HMI tags "DB_SDC_ERROR_STAT_EMS031"
   "DB_SDC_ERRORS_STAT_ER_AKT[31].ER_TRIGER" : Word = PLC DB_SDC_ERRORS_STAT.ER_AKT[31].ER_TRIGER AT %DB3724.DBW30000, 1 s
   "DB_SDC_ERRORS_STAT_ER_AKT[31].ER_STAT[1].DRIVE_POS" : DInt = PLC DB_SDC_ERRORS_STAT.ER_AKT[31].ER_STAT[1].DRIVE_POS AT %DB3724.DBD30006, 1 s
   "DB_SDC_ERRORS_STAT_ER_AKT[31].ER_STAT[1].ERROR" : Int = PLC DB_SDC_ERRORS_STAT.ER_AKT[31].ER_STAT[1].ERROR AT %DB3724.DBW30012, 1 s
   "DB_SDC_ERRORS_STAT_ER_AKT[31].ER_STAT[2].DRIVE_POS" : DInt = PLC DB_SDC_ERRORS_STAT.ER_AKT[31].ER_STAT[2].DRIVE_POS AT %DB3724.DBD30022, 1 s
   "DB_SDC_ERRORS_STAT_ER_AKT[31].ER_STAT[2].ERROR" : Int = PLC DB_SDC_ERRORS_STAT.ER_AKT[31].ER_STAT[2].ERROR AT %DB3724.DBW30028, 1 s
   "DB_SDC_ERRORS_STAT_ER_AKT[31].ER_STAT[3].DRIVE_POS" : DInt = PLC DB_SDC_ERRORS_STAT.ER_AKT[31].ER_STAT[3].DRIVE_POS AT %DB3724.DBD30038, 1 s
   "DB_SDC_ERRORS_STAT_ER_AKT[31].ER_STAT[3].ERROR" : Int = PLC DB_SDC_ERRORS_STAT.ER_AKT[31].ER_STAT[3].ERROR AT %DB3724.DBW30044, 1 s
   "DB_SDC_ERRORS_STAT_ER_AKT[31].ER_STAT[4].DRIVE_POS" : DInt = PLC DB_SDC_ERRORS_STAT.ER_AKT[31].ER_STAT[4].DRIVE_POS AT %DB3724.DBD30054, 1 s
   "DB_SDC_ERRORS_STAT_ER_AKT[31].ER_STAT[4].ERROR" : Int = PLC DB_SDC_ERRORS_STAT.ER_AKT[31].ER_STAT[4].ERROR AT %DB3724.DBW30060, 1 s

HMI tags "DB_SDC_ERROR_STAT_EMS032"
   "DB_SDC_ERRORS_STAT_ER_AKT[32].ER_TRIGER" : Word = PLC DB_SDC_ERRORS_STAT.ER_AKT[32].ER_TRIGER AT %DB3724.DBW30066, 1 s
   "DB_SDC_ERRORS_STAT_ER_AKT[32].ER_STAT[1].DRIVE_POS" : DInt = PLC DB_SDC_ERRORS_STAT.ER_AKT[32].ER_STAT[1].DRIVE_POS AT %DB3724.DBD30072, 1 s
   "DB_SDC_ERRORS_STAT_ER_AKT[32].ER_STAT[1].ERROR" : Int = PLC DB_SDC_ERRORS_STAT.ER_AKT[32].ER_STAT[1].ERROR AT %DB3724.DBW30078, 1 s
   "DB_SDC_ERRORS_STAT_ER_AKT[32].ER_STAT[2].DRIVE_POS" : DInt = PLC DB_SDC_ERRORS_STAT.ER_AKT[32].ER_STAT[2].DRIVE_POS AT %DB3724.DBD30088, 1 s
   "DB_SDC_ERRORS_STAT_ER_AKT[32].ER_STAT[2].ERROR" : Int = PLC DB_SDC_ERRORS_STAT.ER_AKT[32].ER_STAT[2].ERROR AT %DB3724.DBW30094, 1 s
   "DB_SDC_ERRORS_STAT_ER_AKT[32].ER_STAT[3].DRIVE_POS" : DInt = PLC DB_SDC_ERRORS_STAT.ER_AKT[32].ER_STAT[3].DRIVE_POS AT %DB3724.DBD30104, 1 s
   "DB_SDC_ERRORS_STAT_ER_AKT[32].ER_STAT[3].ERROR" : Int = PLC DB_SDC_ERRORS_STAT.ER_AKT[32].ER_STAT[3].ERROR AT %DB3724.DBW30110, 1 s
   "DB_SDC_ERRORS_STAT_ER_AKT[32].ER_STAT[4].DRIVE_POS" : DInt = PLC DB_SDC_ERRORS_STAT.ER_AKT[32].ER_STAT[4].DRIVE_POS AT %DB3724.DBD30120, 1 s
   "DB_SDC_ERRORS_STAT_ER_AKT[32].ER_STAT[4].ERROR" : Int = PLC DB_SDC_ERRORS_STAT.ER_AKT[32].ER_STAT[4].ERROR AT %DB3724.DBW30126, 1 s

HMI tags "DB_SDC_ERROR_STAT_EMS033"
   "DB_SDC_ERRORS_STAT_ER_AKT[33].ER_TRIGER" : Word = PLC DB_SDC_ERRORS_STAT.ER_AKT[33].ER_TRIGER AT %DB3724.DBW30132, 1 s
   "DB_SDC_ERRORS_STAT_ER_AKT[33].ER_STAT[1].DRIVE_POS" : DInt = PLC DB_SDC_ERRORS_STAT.ER_AKT[33].ER_STAT[1].DRIVE_POS AT %DB3724.DBD30138, 1 s
   "DB_SDC_ERRORS_STAT_ER_AKT[33].ER_STAT[1].ERROR" : Int = PLC DB_SDC_ERRORS_STAT.ER_AKT[33].ER_STAT[1].ERROR AT %DB3724.DBW30144, 1 s
   "DB_SDC_ERRORS_STAT_ER_AKT[33].ER_STAT[2].DRIVE_POS" : DInt = PLC DB_SDC_ERRORS_STAT.ER_AKT[63].ER_STAT[4].DRIVE_POS AT %DB3724.DBD30154, 1 s
   "DB_SDC_ERRORS_STAT_ER_AKT[33].ER_STAT[2].ERROR" : Int = PLC DB_SDC_ERRORS_STAT.ER_AKT[33].ER_STAT[2].ERROR AT %DB3724.DBW30160, 1 s
   "DB_SDC_ERRORS_STAT_ER_AKT[33].ER_STAT[3].DRIVE_POS" : DInt = PLC DB_SDC_ERRORS_STAT.ER_AKT[33].ER_STAT[3].DRIVE_POS AT %DB3724.DBD30170, 1 s
   "DB_SDC_ERRORS_STAT_ER_AKT[33].ER_STAT[3].ERROR" : Int = PLC DB_SDC_ERRORS_STAT.ER_AKT[33].ER_STAT[3].ERROR AT %DB3724.DBW30176, 1 s
   "DB_SDC_ERRORS_STAT_ER_AKT[33].ER_STAT[4].DRIVE_POS" : DInt = PLC DB_SDC_ERRORS_STAT.ER_AKT[33].ER_STAT[4].DRIVE_POS AT %DB3724.DBD30186, 1 s
   "DB_SDC_ERRORS_STAT_ER_AKT[33].ER_STAT[4].ERROR" : Int = PLC DB_SDC_ERRORS_STAT.ER_AKT[33].ER_STAT[4].ERROR AT %DB3724.DBW30192, 1 s

HMI tags "DB_SDC_ERROR_STAT_EMS034"
   "DB_SDC_ERRORS_STAT_ER_AKT[34].ER_TRIGER" : Word = PLC DB_SDC_ERRORS_STAT.ER_AKT[34].ER_TRIGER AT %DB3724.DBW30198, 1 s
   "DB_SDC_ERRORS_STAT_ER_AKT[34].ER_STAT[1].DRIVE_POS" : DInt = PLC DB_SDC_ERRORS_STAT.ER_AKT[34].ER_STAT[1].DRIVE_POS AT %DB3724.DBD30204, 1 s
   "DB_SDC_ERRORS_STAT_ER_AKT[34].ER_STAT[1].ERROR" : Int = PLC DB_SDC_ERRORS_STAT.ER_AKT[34].ER_STAT[1].ERROR AT %DB3724.DBW30210, 1 s
   "DB_SDC_ERRORS_STAT_ER_AKT[34].ER_STAT[2].DRIVE_POS" : DInt = PLC DB_SDC_ERRORS_STAT.ER_AKT[34].ER_STAT[2].DRIVE_POS AT %DB3724.DBD30220, 1 s
   "DB_SDC_ERRORS_STAT_ER_AKT[34].ER_STAT[2].ERROR" : Int = PLC DB_SDC_ERRORS_STAT.ER_AKT[34].ER_STAT[2].ERROR AT %DB3724.DBW30226, 1 s
   "DB_SDC_ERRORS_STAT_ER_AKT[34].ER_STAT[3].DRIVE_POS" : DInt = PLC DB_SDC_ERRORS_STAT.ER_AKT[34].ER_STAT[3].DRIVE_POS AT %DB3724.DBD30236, 1 s
   "DB_SDC_ERRORS_STAT_ER_AKT[34].ER_STAT[3].ERROR" : Int = PLC DB_SDC_ERRORS_STAT.ER_AKT[34].ER_STAT[3].ERROR AT %DB3724.DBW30242, 1 s
   "DB_SDC_ERRORS_STAT_ER_AKT[34].ER_STAT[4].DRIVE_POS" : DInt = PLC DB_SDC_ERRORS_STAT.ER_AKT[34].ER_STAT[4].DRIVE_POS AT %DB3724.DBD30252, 1 s
   "DB_SDC_ERRORS_STAT_ER_AKT[34].ER_STAT[4].ERROR" : Int = PLC DB_SDC_ERRORS_STAT.ER_AKT[34].ER_STAT[4].ERROR AT %DB3724.DBW30258, 1 s

HMI tags "DB_SDC_ERROR_STAT_EMS035"
   "DB_SDC_ERRORS_STAT_ER_AKT[35].ER_TRIGER" : Word = PLC DB_SDC_ERRORS_STAT.ER_AKT[35].ER_TRIGER AT %DB3724.DBW30264, 1 s
   "DB_SDC_ERRORS_STAT_ER_AKT[35].ER_STAT[1].DRIVE_POS" : DInt = PLC DB_SDC_ERRORS_STAT.ER_AKT[35].ER_STAT[1].DRIVE_POS AT %DB3724.DBD30270, 1 s
   "DB_SDC_ERRORS_STAT_ER_AKT[35].ER_STAT[1].ERROR" : Int = PLC DB_SDC_ERRORS_STAT.ER_AKT[35].ER_STAT[1].ERROR AT %DB3724.DBW30276, 1 s
   "DB_SDC_ERRORS_STAT_ER_AKT[35].ER_STAT[2].DRIVE_POS" : DInt = PLC DB_SDC_ERRORS_STAT.ER_AKT[35].ER_STAT[2].DRIVE_POS AT %DB3724.DBD30286, 1 s
   "DB_SDC_ERRORS_STAT_ER_AKT[35].ER_STAT[2].ERROR" : Int = PLC DB_SDC_ERRORS_STAT.ER_AKT[35].ER_STAT[2].ERROR AT %DB3724.DBW30292, 1 s
   "DB_SDC_ERRORS_STAT_ER_AKT[35].ER_STAT[3].DRIVE_POS" : DInt = PLC DB_SDC_ERRORS_STAT.ER_AKT[35].ER_STAT[3].DRIVE_POS AT %DB3724.DBD30302, 1 s
   "DB_SDC_ERRORS_STAT_ER_AKT[35].ER_STAT[3].ERROR" : Int = PLC DB_SDC_ERRORS_STAT.ER_AKT[35].ER_STAT[3].ERROR AT %DB3724.DBW30308, 1 s
   "DB_SDC_ERRORS_STAT_ER_AKT[35].ER_STAT[4].DRIVE_POS" : DInt = PLC DB_SDC_ERRORS_STAT.ER_AKT[35].ER_STAT[4].DRIVE_POS AT %DB3724.DBD30318, 1 s
   "DB_SDC_ERRORS_STAT_ER_AKT[35].ER_STAT[4].ERROR" : Int = PLC DB_SDC_ERRORS_STAT.ER_AKT[35].ER_STAT[4].ERROR AT %DB3724.DBW30324, 1 s

HMI tags "DB_SDC_ERROR_STAT_EMS036"
   "DB_SDC_ERRORS_STAT_ER_AKT[36].ER_TRIGER" : Word = PLC DB_SDC_ERRORS_STAT.ER_AKT[36].ER_TRIGER AT %DB3724.DBW30330, 1 s
   "DB_SDC_ERRORS_STAT_ER_AKT[36].ER_STAT[1].DRIVE_POS" : DInt = PLC DB_SDC_ERRORS_STAT.ER_AKT[36].ER_STAT[1].DRIVE_POS AT %DB3724.DBD30336, 1 s
   "DB_SDC_ERRORS_STAT_ER_AKT[36].ER_STAT[1].ERROR" : Int = PLC DB_SDC_ERRORS_STAT.ER_AKT[36].ER_STAT[1].ERROR AT %DB3724.DBW30342, 1 s
   "DB_SDC_ERRORS_STAT_ER_AKT[36].ER_STAT[2].DRIVE_POS" : DInt = PLC DB_SDC_ERRORS_STAT.ER_AKT[36].ER_STAT[2].DRIVE_POS AT %DB3724.DBD30352, 1 s
   "DB_SDC_ERRORS_STAT_ER_AKT[36].ER_STAT[2].ERROR" : Int = PLC DB_SDC_ERRORS_STAT.ER_AKT[36].ER_STAT[2].ERROR AT %DB3724.DBW30358, 1 s
   "DB_SDC_ERRORS_STAT_ER_AKT[36].ER_STAT[3].DRIVE_POS" : DInt = PLC DB_SDC_ERRORS_STAT.ER_AKT[36].ER_STAT[3].DRIVE_POS AT %DB3724.DBD30368, 1 s
   "DB_SDC_ERRORS_STAT_ER_AKT[36].ER_STAT[3].ERROR" : Int = PLC DB_SDC_ERRORS_STAT.ER_AKT[36].ER_STAT[3].ERROR AT %DB3724.DBW30374, 1 s
   "DB_SDC_ERRORS_STAT_ER_AKT[36].ER_STAT[4].DRIVE_POS" : DInt = PLC DB_SDC_ERRORS_STAT.ER_AKT[36].ER_STAT[4].DRIVE_POS AT %DB3724.DBD30384, 1 s
   "DB_SDC_ERRORS_STAT_ER_AKT[36].ER_STAT[4].ERROR" : Int = PLC DB_SDC_ERRORS_STAT.ER_AKT[36].ER_STAT[4].ERROR AT %DB3724.DBW30390, 1 s

HMI tags "DB_SDC_ERROR_STAT_EMS037"
   "DB_SDC_ERRORS_STAT_ER_AKT[37].ER_TRIGER" : Word = PLC DB_SDC_ERRORS_STAT.ER_AKT[37].ER_TRIGER AT %DB3724.DBW30396, 1 s
   "DB_SDC_ERRORS_STAT_ER_AKT[37].ER_STAT[1].DRIVE_POS" : DInt = PLC DB_SDC_ERRORS_STAT.ER_AKT[37].ER_STAT[1].DRIVE_POS AT %DB3724.DBD30402, 1 s
   "DB_SDC_ERRORS_STAT_ER_AKT[37].ER_STAT[1].ERROR" : Int = PLC DB_SDC_ERRORS_STAT.ER_AKT[37].ER_STAT[1].ERROR AT %DB3724.DBW30408, 1 s
   "DB_SDC_ERRORS_STAT_ER_AKT[37].ER_STAT[2].DRIVE_POS" : DInt = PLC DB_SDC_ERRORS_STAT.ER_AKT[37].ER_STAT[2].DRIVE_POS AT %DB3724.DBD30418, 1 s
   "DB_SDC_ERRORS_STAT_ER_AKT[37].ER_STAT[2].ERROR" : Int = PLC DB_SDC_ERRORS_STAT.ER_AKT[37].ER_STAT[2].ERROR AT %DB3724.DBW30424, 1 s
   "DB_SDC_ERRORS_STAT_ER_AKT[37].ER_STAT[3].DRIVE_POS" : DInt = PLC DB_SDC_ERRORS_STAT.ER_AKT[37].ER_STAT[3].DRIVE_POS AT %DB3724.DBD30434, 1 s
   "DB_SDC_ERRORS_STAT_ER_AKT[37].ER_STAT[3].ERROR" : Int = PLC DB_SDC_ERRORS_STAT.ER_AKT[37].ER_STAT[3].ERROR AT %DB3724.DBW30440, 1 s
   "DB_SDC_ERRORS_STAT_ER_AKT[37].ER_STAT[4].DRIVE_POS" : DInt = PLC DB_SDC_ERRORS_STAT.ER_AKT[37].ER_STAT[4].DRIVE_POS AT %DB3724.DBD30450, 1 s
   "DB_SDC_ERRORS_STAT_ER_AKT[37].ER_STAT[4].ERROR" : Int = PLC DB_SDC_ERRORS_STAT.ER_AKT[37].ER_STAT[4].ERROR AT %DB3724.DBW30456, 1 s

HMI tags "DB_SDC_ERROR_STAT_EMS038"
   "DB_SDC_ERRORS_STAT_ER_AKT[38].ER_TRIGER" : Word = PLC DB_SDC_ERRORS_STAT.ER_AKT[38].ER_TRIGER AT %DB3724.DBW30462, 1 s
   "DB_SDC_ERRORS_STAT_ER_AKT[38].ER_STAT[1].DRIVE_POS" : DInt = PLC DB_SDC_ERRORS_STAT.ER_AKT[38].ER_STAT[1].DRIVE_POS AT %DB3724.DBD30468, 1 s
   "DB_SDC_ERRORS_STAT_ER_AKT[38].ER_STAT[1].ERROR" : Int = PLC DB_SDC_ERRORS_STAT.ER_AKT[38].ER_STAT[1].ERROR AT %DB3724.DBW30474, 1 s
   "DB_SDC_ERRORS_STAT_ER_AKT[38].ER_STAT[2].DRIVE_POS" : DInt = PLC DB_SDC_ERRORS_STAT.ER_AKT[38].ER_STAT[2].DRIVE_POS AT %DB3724.DBD30484, 1 s
   "DB_SDC_ERRORS_STAT_ER_AKT[38].ER_STAT[2].ERROR" : Int = PLC DB_SDC_ERRORS_STAT.ER_AKT[38].ER_STAT[2].ERROR AT %DB3724.DBW30490, 1 s
   "DB_SDC_ERRORS_STAT_ER_AKT[38].ER_STAT[3].DRIVE_POS" : DInt = PLC DB_SDC_ERRORS_STAT.ER_AKT[38].ER_STAT[3].DRIVE_POS AT %DB3724.DBD30500, 1 s
   "DB_SDC_ERRORS_STAT_ER_AKT[38].ER_STAT[3].ERROR" : Int = PLC DB_SDC_ERRORS_STAT.ER_AKT[38].ER_STAT[3].ERROR AT %DB3724.DBW30506, 1 s
   "DB_SDC_ERRORS_STAT_ER_AKT[38].ER_STAT[4].DRIVE_POS" : DInt = PLC DB_SDC_ERRORS_STAT.ER_AKT[38].ER_STAT[4].DRIVE_POS AT %DB3724.DBD30516, 1 s
   "DB_SDC_ERRORS_STAT_ER_AKT[38].ER_STAT[4].ERROR" : Int = PLC DB_SDC_ERRORS_STAT.ER_AKT[38].ER_STAT[4].ERROR AT %DB3724.DBW30522, 1 s

HMI tags "DB_SDC_ERROR_STAT_EMS039"
   "DB_SDC_ERRORS_STAT_ER_AKT[39].ER_TRIGER" : Word = PLC DB_SDC_ERRORS_STAT.ER_AKT[39].ER_TRIGER AT %DB3724.DBW30528, 1 s
   "DB_SDC_ERRORS_STAT_ER_AKT[39].ER_STAT[1].DRIVE_POS" : DInt = PLC DB_SDC_ERRORS_STAT.ER_AKT[39].ER_STAT[1].DRIVE_POS AT %DB3724.DBD30534, 1 s
   "DB_SDC_ERRORS_STAT_ER_AKT[39].ER_STAT[1].ERROR" : Int = PLC DB_SDC_ERRORS_STAT.ER_AKT[39].ER_STAT[1].ERROR AT %DB3724.DBW30540, 1 s
   "DB_SDC_ERRORS_STAT_ER_AKT[39].ER_STAT[2].DRIVE_POS" : DInt = PLC DB_SDC_ERRORS_STAT.ER_AKT[39].ER_STAT[2].DRIVE_POS AT %DB3724.DBD30550, 1 s
   "DB_SDC_ERRORS_STAT_ER_AKT[39].ER_STAT[2].ERROR" : Int = PLC DB_SDC_ERRORS_STAT.ER_AKT[39].ER_STAT[2].ERROR AT %DB3724.DBW30556, 1 s
   "DB_SDC_ERRORS_STAT_ER_AKT[39].ER_STAT[3].DRIVE_POS" : DInt = PLC DB_SDC_ERRORS_STAT.ER_AKT[39].ER_STAT[3].DRIVE_POS AT %DB3724.DBD30566, 1 s
   "DB_SDC_ERRORS_STAT_ER_AKT[39].ER_STAT[3].ERROR" : Int = PLC DB_SDC_ERRORS_STAT.ER_AKT[39].ER_STAT[3].ERROR AT %DB3724.DBW30572, 1 s
   "DB_SDC_ERRORS_STAT_ER_AKT[39].ER_STAT[4].DRIVE_POS" : DInt = PLC DB_SDC_ERRORS_STAT.ER_AKT[39].ER_STAT[4].DRIVE_POS AT %DB3724.DBD30582, 1 s
   "DB_SDC_ERRORS_STAT_ER_AKT[39].ER_STAT[4].ERROR" : Int = PLC DB_SDC_ERRORS_STAT.ER_AKT[39].ER_STAT[4].ERROR AT %DB3724.DBW30588, 1 s

HMI tags "DB_SDC_ERROR_STAT_EMS040"
   "DB_SDC_ERRORS_STAT_ER_AKT[40].ER_TRIGER" : Word = PLC DB_SDC_ERRORS_STAT.ER_AKT[40].ER_TRIGER AT %DB3724.DBW30594, 1 s
   "DB_SDC_ERRORS_STAT_ER_AKT[40].ER_STAT[1].DRIVE_POS" : DInt = PLC DB_SDC_ERRORS_STAT.ER_AKT[40].ER_STAT[1].DRIVE_POS AT %DB3724.DBD30600, 1 s
   "DB_SDC_ERRORS_STAT_ER_AKT[40].ER_STAT[1].ERROR" : Int = PLC DB_SDC_ERRORS_STAT.ER_AKT[40].ER_STAT[1].ERROR AT %DB3724.DBW30606, 1 s
   "DB_SDC_ERRORS_STAT_ER_AKT[40].ER_STAT[2].DRIVE_POS" : DInt = PLC DB_SDC_ERRORS_STAT.ER_AKT[40].ER_STAT[2].DRIVE_POS AT %DB3724.DBD30616, 1 s
   "DB_SDC_ERRORS_STAT_ER_AKT[40].ER_STAT[2].ERROR" : Int = PLC DB_SDC_ERRORS_STAT.ER_AKT[40].ER_STAT[2].ERROR AT %DB3724.DBW30622, 1 s
   "DB_SDC_ERRORS_STAT_ER_AKT[40].ER_STAT[3].DRIVE_POS" : DInt = PLC DB_SDC_ERRORS_STAT.ER_AKT[40].ER_STAT[3].DRIVE_POS AT %DB3724.DBD30632, 1 s
   "DB_SDC_ERRORS_STAT_ER_AKT[40].ER_STAT[3].ERROR" : Int = PLC DB_SDC_ERRORS_STAT.ER_AKT[40].ER_STAT[3].ERROR AT %DB3724.DBW30638, 1 s
   "DB_SDC_ERRORS_STAT_ER_AKT[40].ER_STAT[4].DRIVE_POS" : DInt = PLC DB_SDC_ERRORS_STAT.ER_AKT[40].ER_STAT[4].DRIVE_POS AT %DB3724.DBD30648, 1 s
   "DB_SDC_ERRORS_STAT_ER_AKT[40].ER_STAT[4].ERROR" : Int = PLC DB_SDC_ERRORS_STAT.ER_AKT[40].ER_STAT[4].ERROR AT %DB3724.DBW30654, 1 s

HMI tags "DB_SDC_ERROR_STAT_EMS041"
   "DB_SDC_ERRORS_STAT_ER_AKT[41].ER_TRIGER" : Word = PLC DB_SDC_ERRORS_STAT.ER_AKT[41].ER_TRIGER AT %DB3724.DBW30660, 1 s
   "DB_SDC_ERRORS_STAT_ER_AKT[41].ER_STAT[1].DRIVE_POS" : DInt = PLC DB_SDC_ERRORS_STAT.ER_AKT[41].ER_STAT[1].DRIVE_POS AT %DB3724.DBD30666, 1 s
   "DB_SDC_ERRORS_STAT_ER_AKT[41].ER_STAT[1].ERROR" : Int = PLC DB_SDC_ERRORS_STAT.ER_AKT[41].ER_STAT[1].ERROR AT %DB3724.DBW30672, 1 s
   "DB_SDC_ERRORS_STAT_ER_AKT[41].ER_STAT[2].DRIVE_POS" : DInt = PLC DB_SDC_ERRORS_STAT.ER_AKT[41].ER_STAT[2].DRIVE_POS AT %DB3724.DBD30682, 1 s
   "DB_SDC_ERRORS_STAT_ER_AKT[41].ER_STAT[2].ERROR" : Int = PLC DB_SDC_ERRORS_STAT.ER_AKT[41].ER_STAT[2].ERROR AT %DB3724.DBW30688, 1 s
   "DB_SDC_ERRORS_STAT_ER_AKT[41].ER_STAT[3].DRIVE_POS" : DInt = PLC DB_SDC_ERRORS_STAT.ER_AKT[41].ER_STAT[3].DRIVE_POS AT %DB3724.DBD30698, 1 s
   "DB_SDC_ERRORS_STAT_ER_AKT[41].ER_STAT[3].ERROR" : Int = PLC DB_SDC_ERRORS_STAT.ER_AKT[41].ER_STAT[3].ERROR AT %DB3724.DBW30704, 1 s
   "DB_SDC_ERRORS_STAT_ER_AKT[41].ER_STAT[4].DRIVE_POS" : DInt = PLC DB_SDC_ERRORS_STAT.ER_AKT[41].ER_STAT[4].DRIVE_POS AT %DB3724.DBD30714, 1 s
   "DB_SDC_ERRORS_STAT_ER_AKT[41].ER_STAT[4].ERROR" : Int = PLC DB_SDC_ERRORS_STAT.ER_AKT[41].ER_STAT[4].ERROR AT %DB3724.DBW30720, 1 s

HMI tags "DB_SDC_ERROR_STAT_EMS042"
   "DB_SDC_ERRORS_STAT_ER_AKT[42].ER_TRIGER" : Word = PLC DB_SDC_ERRORS_STAT.ER_AKT[42].ER_TRIGER AT %DB3724.DBW30726, 1 s
   "DB_SDC_ERRORS_STAT_ER_AKT[42].ER_STAT[1].DRIVE_POS" : DInt = PLC DB_SDC_ERRORS_STAT.ER_AKT[42].ER_STAT[1].DRIVE_POS AT %DB3724.DBD30732, 1 s
   "DB_SDC_ERRORS_STAT_ER_AKT[42].ER_STAT[1].ERROR" : Int = PLC DB_SDC_ERRORS_STAT.ER_AKT[42].ER_STAT[1].ERROR AT %DB3724.DBW30738, 1 s
   "DB_SDC_ERRORS_STAT_ER_AKT[42].ER_STAT[2].DRIVE_POS" : DInt = PLC DB_SDC_ERRORS_STAT.ER_AKT[42].ER_STAT[2].DRIVE_POS AT %DB3724.DBD30748, 1 s
   "DB_SDC_ERRORS_STAT_ER_AKT[42].ER_STAT[2].ERROR" : Int = PLC DB_SDC_ERRORS_STAT.ER_AKT[42].ER_STAT[2].ERROR AT %DB3724.DBW30754, 1 s
   "DB_SDC_ERRORS_STAT_ER_AKT[42].ER_STAT[3].DRIVE_POS" : DInt = PLC DB_SDC_ERRORS_STAT.ER_AKT[42].ER_STAT[3].DRIVE_POS AT %DB3724.DBD30764, 1 s
   "DB_SDC_ERRORS_STAT_ER_AKT[42].ER_STAT[3].ERROR" : Int = PLC DB_SDC_ERRORS_STAT.ER_AKT[42].ER_STAT[3].ERROR AT %DB3724.DBW30770, 1 s
   "DB_SDC_ERRORS_STAT_ER_AKT[42].ER_STAT[4].DRIVE_POS" : DInt = PLC DB_SDC_ERRORS_STAT.ER_AKT[42].ER_STAT[4].DRIVE_POS AT %DB3724.DBD30780, 1 s
   "DB_SDC_ERRORS_STAT_ER_AKT[42].ER_STAT[4].ERROR" : Int = PLC DB_SDC_ERRORS_STAT.ER_AKT[42].ER_STAT[4].ERROR AT %DB3724.DBW30786, 1 s

HMI tags "DB_SDC_ERROR_STAT_EMS043"
   "DB_SDC_ERRORS_STAT_ER_AKT[43].ER_TRIGER" : Word = PLC DB_SDC_ERRORS_STAT.ER_AKT[43].ER_TRIGER AT %DB3724.DBW30792, 1 s
   "DB_SDC_ERRORS_STAT_ER_AKT[43].ER_STAT[1].DRIVE_POS" : DInt = PLC DB_SDC_ERRORS_STAT.ER_AKT[43].ER_STAT[1].DRIVE_POS AT %DB3724.DBD30798, 1 s
   "DB_SDC_ERRORS_STAT_ER_AKT[43].ER_STAT[1].ERROR" : Int = PLC DB_SDC_ERRORS_STAT.ER_AKT[43].ER_STAT[1].ERROR AT %DB3724.DBW30804, 1 s
   "DB_SDC_ERRORS_STAT_ER_AKT[43].ER_STAT[2].DRIVE_POS" : DInt = PLC DB_SDC_ERRORS_STAT.ER_AKT[43].ER_STAT[2].DRIVE_POS AT %DB3724.DBD30814, 1 s
   "DB_SDC_ERRORS_STAT_ER_AKT[43].ER_STAT[2].ERROR" : Int = PLC DB_SDC_ERRORS_STAT.ER_AKT[43].ER_STAT[2].ERROR AT %DB3724.DBW30820, 1 s
   "DB_SDC_ERRORS_STAT_ER_AKT[43].ER_STAT[3].DRIVE_POS" : DInt = PLC DB_SDC_ERRORS_STAT.ER_AKT[43].ER_STAT[3].DRIVE_POS AT %DB3724.DBD30830, 1 s
   "DB_SDC_ERRORS_STAT_ER_AKT[43].ER_STAT[3].ERROR" : Int = PLC DB_SDC_ERRORS_STAT.ER_AKT[43].ER_STAT[3].ERROR AT %DB3724.DBW30836, 1 s
   "DB_SDC_ERRORS_STAT_ER_AKT[43].ER_STAT[4].DRIVE_POS" : DInt = PLC DB_SDC_ERRORS_STAT.ER_AKT[43].ER_STAT[4].DRIVE_POS AT %DB3724.DBD30846, 1 s
   "DB_SDC_ERRORS_STAT_ER_AKT[43].ER_STAT[4].ERROR" : Int = PLC DB_SDC_ERRORS_STAT.ER_AKT[43].ER_STAT[4].ERROR AT %DB3724.DBW30852, 1 s

HMI tags "DB_SDC_ERROR_STAT_EMS044"
   "DB_SDC_ERRORS_STAT_ER_AKT[44].ER_TRIGER" : Word = PLC DB_SDC_ERRORS_STAT.ER_AKT[44].ER_TRIGER AT %DB3724.DBW30858, 1 s
   "DB_SDC_ERRORS_STAT_ER_AKT[44].ER_STAT[1].DRIVE_POS" : DInt = PLC DB_SDC_ERRORS_STAT.ER_AKT[44].ER_STAT[1].DRIVE_POS AT %DB3724.DBD30864, 1 s
   "DB_SDC_ERRORS_STAT_ER_AKT[44].ER_STAT[1].ERROR" : Int = PLC DB_SDC_ERRORS_STAT.ER_AKT[44].ER_STAT[1].ERROR AT %DB3724.DBW30870, 1 s
   "DB_SDC_ERRORS_STAT_ER_AKT[44].ER_STAT[2].DRIVE_POS" : DInt = PLC DB_SDC_ERRORS_STAT.ER_AKT[44].ER_STAT[2].DRIVE_POS AT %DB3724.DBD30880, 1 s
   "DB_SDC_ERRORS_STAT_ER_AKT[44].ER_STAT[2].ERROR" : Int = PLC DB_SDC_ERRORS_STAT.ER_AKT[44].ER_STAT[2].ERROR AT %DB3724.DBW30886, 1 s
   "DB_SDC_ERRORS_STAT_ER_AKT[44].ER_STAT[3].DRIVE_POS" : DInt = PLC DB_SDC_ERRORS_STAT.ER_AKT[44].ER_STAT[3].DRIVE_POS AT %DB3724.DBD30896, 1 s
   "DB_SDC_ERRORS_STAT_ER_AKT[44].ER_STAT[3].ERROR" : Int = PLC DB_SDC_ERRORS_STAT.ER_AKT[44].ER_STAT[3].ERROR AT %DB3724.DBW30902, 1 s
   "DB_SDC_ERRORS_STAT_ER_AKT[44].ER_STAT[4].DRIVE_POS" : DInt = PLC DB_SDC_ERRORS_STAT.ER_AKT[44].ER_STAT[4].DRIVE_POS AT %DB3724.DBD30912, 1 s
   "DB_SDC_ERRORS_STAT_ER_AKT[44].ER_STAT[4].ERROR" : Int = PLC DB_SDC_ERRORS_STAT.ER_AKT[44].ER_STAT[4].ERROR AT %DB3724.DBW30918, 1 s

HMI tags "DB_SDC_ERROR_STAT_EMS045"
   "DB_SDC_ERRORS_STAT_ER_AKT[45].ER_TRIGER" : Word = PLC DB_SDC_ERRORS_STAT.ER_AKT[45].ER_TRIGER AT %DB3724.DBW30924, 1 s
   "DB_SDC_ERRORS_STAT_ER_AKT[45].ER_STAT[1].DRIVE_POS" : DInt = PLC DB_SDC_ERRORS_STAT.ER_AKT[45].ER_STAT[1].DRIVE_POS AT %DB3724.DBD30930, 1 s
   "DB_SDC_ERRORS_STAT_ER_AKT[45].ER_STAT[1].ERROR" : Int = PLC DB_SDC_ERRORS_STAT.ER_AKT[45].ER_STAT[1].ERROR AT %DB3724.DBW30936, 1 s
   "DB_SDC_ERRORS_STAT_ER_AKT[45].ER_STAT[2].DRIVE_POS" : DInt = PLC DB_SDC_ERRORS_STAT.ER_AKT[45].ER_STAT[2].DRIVE_POS AT %DB3724.DBD30946, 1 s
   "DB_SDC_ERRORS_STAT_ER_AKT[45].ER_STAT[2].ERROR" : Int = PLC DB_SDC_ERRORS_STAT.ER_AKT[45].ER_STAT[2].ERROR AT %DB3724.DBW30952, 1 s
   "DB_SDC_ERRORS_STAT_ER_AKT[45].ER_STAT[3].DRIVE_POS" : DInt = PLC DB_SDC_ERRORS_STAT.ER_AKT[45].ER_STAT[3].DRIVE_POS AT %DB3724.DBD30962, 1 s
   "DB_SDC_ERRORS_STAT_ER_AKT[45].ER_STAT[3].ERROR" : Int = PLC DB_SDC_ERRORS_STAT.ER_AKT[45].ER_STAT[3].ERROR AT %DB3724.DBW30968, 1 s
   "DB_SDC_ERRORS_STAT_ER_AKT[45].ER_STAT[4].DRIVE_POS" : DInt = PLC DB_SDC_ERRORS_STAT.ER_AKT[45].ER_STAT[4].DRIVE_POS AT %DB3724.DBD30978, 1 s
   "DB_SDC_ERRORS_STAT_ER_AKT[45].ER_STAT[4].ERROR" : Int = PLC DB_SDC_ERRORS_STAT.ER_AKT[45].ER_STAT[4].ERROR AT %DB3724.DBW30984, 1 s

HMI tags "DB_SDC_ERROR_STAT_EMS046"
   "DB_SDC_ERRORS_STAT_ER_AKT[46].ER_TRIGER" : Word = PLC DB_SDC_ERRORS_STAT.ER_AKT[46].ER_TRIGER AT %DB3724.DBW30990, 1 s
   "DB_SDC_ERRORS_STAT_ER_AKT[46].ER_STAT[1].DRIVE_POS" : DInt = PLC DB_SDC_ERRORS_STAT.ER_AKT[46].ER_STAT[1].DRIVE_POS AT %DB3724.DBD30996, 1 s
   "DB_SDC_ERRORS_STAT_ER_AKT[46].ER_STAT[1].ERROR" : Int = PLC DB_SDC_ERRORS_STAT.ER_AKT[46].ER_STAT[1].ERROR AT %DB3724.DBW31002, 1 s
   "DB_SDC_ERRORS_STAT_ER_AKT[46].ER_STAT[2].DRIVE_POS" : DInt = PLC DB_SDC_ERRORS_STAT.ER_AKT[46].ER_STAT[2].DRIVE_POS AT %DB3724.DBD31012, 1 s
   "DB_SDC_ERRORS_STAT_ER_AKT[46].ER_STAT[2].ERROR" : Int = PLC DB_SDC_ERRORS_STAT.ER_AKT[46].ER_STAT[2].ERROR AT %DB3724.DBW31018, 1 s
   "DB_SDC_ERRORS_STAT_ER_AKT[46].ER_STAT[3].DRIVE_POS" : DInt = PLC DB_SDC_ERRORS_STAT.ER_AKT[46].ER_STAT[3].DRIVE_POS AT %DB3724.DBD31028, 1 s
   "DB_SDC_ERRORS_STAT_ER_AKT[46].ER_STAT[3].ERROR" : Int = PLC DB_SDC_ERRORS_STAT.ER_AKT[46].ER_STAT[3].ERROR AT %DB3724.DBW31034, 1 s
   "DB_SDC_ERRORS_STAT_ER_AKT[46].ER_STAT[4].DRIVE_POS" : DInt = PLC DB_SDC_ERRORS_STAT.ER_AKT[46].ER_STAT[4].DRIVE_POS AT %DB3724.DBD31044, 1 s
   "DB_SDC_ERRORS_STAT_ER_AKT[46].ER_STAT[4].ERROR" : Int = PLC DB_SDC_ERRORS_STAT.ER_AKT[46].ER_STAT[4].ERROR AT %DB3724.DBW31050, 1 s

HMI tags "DB_SDC_ERROR_STAT_EMS047"
   "DB_SDC_ERRORS_STAT_ER_AKT[47].ER_TRIGER" : Word = PLC DB_SDC_ERRORS_STAT.ER_AKT[47].ER_TRIGER AT %DB3724.DBW31056, 1 s
   "DB_SDC_ERRORS_STAT_ER_AKT[47].ER_STAT[1].DRIVE_POS" : DInt = PLC DB_SDC_ERRORS_STAT.ER_AKT[47].ER_STAT[1].DRIVE_POS AT %DB3724.DBD31062, 1 s
   "DB_SDC_ERRORS_STAT_ER_AKT[47].ER_STAT[1].ERROR" : Int = PLC DB_SDC_ERRORS_STAT.ER_AKT[47].ER_STAT[1].ERROR AT %DB3724.DBW31068, 1 s
   "DB_SDC_ERRORS_STAT_ER_AKT[47].ER_STAT[2].DRIVE_POS" : DInt = PLC DB_SDC_ERRORS_STAT.ER_AKT[47].ER_STAT[2].DRIVE_POS AT %DB3724.DBD31078, 1 s
   "DB_SDC_ERRORS_STAT_ER_AKT[47].ER_STAT[2].ERROR" : Int = PLC DB_SDC_ERRORS_STAT.ER_AKT[47].ER_STAT[2].ERROR AT %DB3724.DBW31084, 1 s
   "DB_SDC_ERRORS_STAT_ER_AKT[47].ER_STAT[3].DRIVE_POS" : DInt = PLC DB_SDC_ERRORS_STAT.ER_AKT[47].ER_STAT[3].DRIVE_POS AT %DB3724.DBD31094, 1 s
   "DB_SDC_ERRORS_STAT_ER_AKT[47].ER_STAT[3].ERROR" : Int = PLC DB_SDC_ERRORS_STAT.ER_AKT[47].ER_STAT[3].ERROR AT %DB3724.DBW31100, 1 s
   "DB_SDC_ERRORS_STAT_ER_AKT[47].ER_STAT[4].DRIVE_POS" : DInt = PLC DB_SDC_ERRORS_STAT.ER_AKT[47].ER_STAT[4].DRIVE_POS AT %DB3724.DBD31110, 1 s
   "DB_SDC_ERRORS_STAT_ER_AKT[47].ER_STAT[4].ERROR" : Int = PLC DB_SDC_ERRORS_STAT.ER_AKT[47].ER_STAT[4].ERROR AT %DB3724.DBW31116, 1 s

HMI tags "DB_SDC_ERROR_STAT_EMS048"
   "DB_SDC_ERRORS_STAT_ER_AKT[48].ER_TRIGER" : Word = PLC DB_SDC_ERRORS_STAT.ER_AKT[48].ER_TRIGER AT %DB3724.DBW31122, 1 s
   "DB_SDC_ERRORS_STAT_ER_AKT[48].ER_STAT[1].DRIVE_POS" : DInt = PLC DB_SDC_ERRORS_STAT.ER_AKT[48].ER_STAT[1].DRIVE_POS AT %DB3724.DBD31128, 1 s
   "DB_SDC_ERRORS_STAT_ER_AKT[48].ER_STAT[1].ERROR" : Int = PLC DB_SDC_ERRORS_STAT.ER_AKT[48].ER_STAT[1].ERROR AT %DB3724.DBW31134, 1 s
   "DB_SDC_ERRORS_STAT_ER_AKT[48].ER_STAT[2].DRIVE_POS" : DInt = PLC DB_SDC_ERRORS_STAT.ER_AKT[48].ER_STAT[2].DRIVE_POS AT %DB3724.DBD31144, 1 s
   "DB_SDC_ERRORS_STAT_ER_AKT[48].ER_STAT[2].ERROR" : Int = PLC DB_SDC_ERRORS_STAT.ER_AKT[48].ER_STAT[2].ERROR AT %DB3724.DBW31150, 1 s
   "DB_SDC_ERRORS_STAT_ER_AKT[48].ER_STAT[3].DRIVE_POS" : DInt = PLC DB_SDC_ERRORS_STAT.ER_AKT[48].ER_STAT[3].DRIVE_POS AT %DB3724.DBD31160, 1 s
   "DB_SDC_ERRORS_STAT_ER_AKT[48].ER_STAT[3].ERROR" : Int = PLC DB_SDC_ERRORS_STAT.ER_AKT[48].ER_STAT[3].ERROR AT %DB3724.DBW31166, 1 s
   "DB_SDC_ERRORS_STAT_ER_AKT[48].ER_STAT[4].DRIVE_POS" : DInt = PLC DB_SDC_ERRORS_STAT.ER_AKT[48].ER_STAT[4].DRIVE_POS AT %DB3724.DBD31176, 1 s
   "DB_SDC_ERRORS_STAT_ER_AKT[48].ER_STAT[4].ERROR" : Int = PLC DB_SDC_ERRORS_STAT.ER_AKT[48].ER_STAT[4].ERROR AT %DB3724.DBW31182, 1 s

HMI tags "DB_SDC_ERROR_STAT_EMS049"
   "DB_SDC_ERRORS_STAT_ER_AKT[49].ER_TRIGER" : Word = PLC DB_SDC_ERRORS_STAT.ER_AKT[49].ER_TRIGER AT %DB3724.DBW31188, 1 s
   "DB_SDC_ERRORS_STAT_ER_AKT[49].ER_STAT[1].DRIVE_POS" : DInt = PLC DB_SDC_ERRORS_STAT.ER_AKT[49].ER_STAT[1].DRIVE_POS AT %DB3724.DBD31194, 1 s
   "DB_SDC_ERRORS_STAT_ER_AKT[49].ER_STAT[1].ERROR" : Int = PLC DB_SDC_ERRORS_STAT.ER_AKT[49].ER_STAT[1].ERROR AT %DB3724.DBW31200, 1 s
   "DB_SDC_ERRORS_STAT_ER_AKT[49].ER_STAT[2].DRIVE_POS" : DInt = PLC DB_SDC_ERRORS_STAT.ER_AKT[49].ER_STAT[2].DRIVE_POS AT %DB3724.DBD31210, 1 s
   "DB_SDC_ERRORS_STAT_ER_AKT[49].ER_STAT[2].ERROR" : Int = PLC DB_SDC_ERRORS_STAT.ER_AKT[49].ER_STAT[2].ERROR AT %DB3724.DBW31216, 1 s
   "DB_SDC_ERRORS_STAT_ER_AKT[49].ER_STAT[3].DRIVE_POS" : DInt = PLC DB_SDC_ERRORS_STAT.ER_AKT[49].ER_STAT[3].DRIVE_POS AT %DB3724.DBD31226, 1 s
   "DB_SDC_ERRORS_STAT_ER_AKT[49].ER_STAT[3].ERROR" : Int = PLC DB_SDC_ERRORS_STAT.ER_AKT[49].ER_STAT[3].ERROR AT %DB3724.DBW31232, 1 s
   "DB_SDC_ERRORS_STAT_ER_AKT[49].ER_STAT[4].DRIVE_POS" : DInt = PLC DB_SDC_ERRORS_STAT.ER_AKT[49].ER_STAT[4].DRIVE_POS AT %DB3724.DBD31242, 1 s
   "DB_SDC_ERRORS_STAT_ER_AKT[49].ER_STAT[4].ERROR" : Int = PLC DB_SDC_ERRORS_STAT.ER_AKT[49].ER_STAT[4].ERROR AT %DB3724.DBW31248, 1 s

HMI tags "DB_SDC_ERROR_STAT_EMS050"
   "DB_SDC_ERRORS_STAT_ER_AKT[50].ER_TRIGER" : Word = PLC DB_SDC_ERRORS_STAT.ER_AKT[50].ER_TRIGER AT %DB3724.DBW31254, 1 s
   "DB_SDC_ERRORS_STAT_ER_AKT[50].ER_STAT[1].DRIVE_POS" : DInt = PLC DB_SDC_ERRORS_STAT.ER_AKT[50].ER_STAT[1].DRIVE_POS AT %DB3724.DBD31260, 1 s
   "DB_SDC_ERRORS_STAT_ER_AKT[50].ER_STAT[1].ERROR" : Int = PLC DB_SDC_ERRORS_STAT.ER_AKT[50].ER_STAT[1].ERROR AT %DB3724.DBW31266, 1 s
   "DB_SDC_ERRORS_STAT_ER_AKT[50].ER_STAT[2].DRIVE_POS" : DInt = PLC DB_SDC_ERRORS_STAT.ER_AKT[50].ER_STAT[2].DRIVE_POS AT %DB3724.DBD31276, 1 s
   "DB_SDC_ERRORS_STAT_ER_AKT[50].ER_STAT[2].ERROR" : Int = PLC DB_SDC_ERRORS_STAT.ER_AKT[50].ER_STAT[2].ERROR AT %DB3724.DBW31282, 1 s
   "DB_SDC_ERRORS_STAT_ER_AKT[50].ER_STAT[3].DRIVE_POS" : DInt = PLC DB_SDC_ERRORS_STAT.ER_AKT[50].ER_STAT[3].DRIVE_POS AT %DB3724.DBD31292, 1 s
   "DB_SDC_ERRORS_STAT_ER_AKT[50].ER_STAT[3].ERROR" : Int = PLC DB_SDC_ERRORS_STAT.ER_AKT[50].ER_STAT[3].ERROR AT %DB3724.DBW31298, 1 s
   "DB_SDC_ERRORS_STAT_ER_AKT[50].ER_STAT[4].DRIVE_POS" : DInt = PLC DB_SDC_ERRORS_STAT.ER_AKT[50].ER_STAT[4].DRIVE_POS AT %DB3724.DBD31308, 1 s
   "DB_SDC_ERRORS_STAT_ER_AKT[50].ER_STAT[4].ERROR" : Int = PLC DB_SDC_ERRORS_STAT.ER_AKT[50].ER_STAT[4].ERROR AT %DB3724.DBW31314, 1 s

HMI tags "DB_SDC_ERROR_STAT_EMS051"
   "DB_SDC_ERRORS_STAT_ER_AKT[51].ER_TRIGER" : Word = PLC DB_SDC_ERRORS_STAT.ER_AKT[51].ER_TRIGER AT %DB3724.DBW31320, 1 s
   "DB_SDC_ERRORS_STAT_ER_AKT[51].ER_STAT[1].DRIVE_POS" : DInt = PLC DB_SDC_ERRORS_STAT.ER_AKT[51].ER_STAT[1].DRIVE_POS AT %DB3724.DBD31326, 1 s
   "DB_SDC_ERRORS_STAT_ER_AKT[51].ER_STAT[1].ERROR" : Int = PLC DB_SDC_ERRORS_STAT.ER_AKT[51].ER_STAT[1].ERROR AT %DB3724.DBW31332, 1 s
   "DB_SDC_ERRORS_STAT_ER_AKT[51].ER_STAT[2].DRIVE_POS" : DInt = PLC DB_SDC_ERRORS_STAT.ER_AKT[51].ER_STAT[2].DRIVE_POS AT %DB3724.DBD31342, 1 s
   "DB_SDC_ERRORS_STAT_ER_AKT[51].ER_STAT[2].ERROR" : Int = PLC DB_SDC_ERRORS_STAT.ER_AKT[51].ER_STAT[2].ERROR AT %DB3724.DBW31348, 1 s
   "DB_SDC_ERRORS_STAT_ER_AKT[51].ER_STAT[3].DRIVE_POS" : DInt = PLC DB_SDC_ERRORS_STAT.ER_AKT[51].ER_STAT[3].DRIVE_POS AT %DB3724.DBD31358, 1 s
   "DB_SDC_ERRORS_STAT_ER_AKT[51].ER_STAT[3].ERROR" : Int = PLC DB_SDC_ERRORS_STAT.ER_AKT[51].ER_STAT[3].ERROR AT %DB3724.DBW31364, 1 s
   "DB_SDC_ERRORS_STAT_ER_AKT[51].ER_STAT[4].DRIVE_POS" : DInt = PLC DB_SDC_ERRORS_STAT.ER_AKT[51].ER_STAT[4].DRIVE_POS AT %DB3724.DBD31374, 1 s
   "DB_SDC_ERRORS_STAT_ER_AKT[51].ER_STAT[4].ERROR" : Int = PLC DB_SDC_ERRORS_STAT.ER_AKT[51].ER_STAT[4].ERROR AT %DB3724.DBW31380, 1 s
